   2165: 'FIT417 1 STARBOARD TANK USD FLOW HIGH', class Tank Control Warnings, trigger "2062_Warning_Data_BTCS_WARNING_WORD_03" bit 5
   2166: 'FIT418 3 PORT TANK USD FLOW LOW', class Tank Control Warnings, trigger "2062_Warning_Data_BTCS_WARNING_WORD_03" bit 6
   2164: 'FIT417 1 STARBOARD TANK USD FLOW LOW', class Tank Control Warnings, trigger "2062_Warning_Data_BTCS_WARNING_WORD_03" bit 4
   2162: 'FIT418 1 PORT TANK USD FLOW LOW', class Tank Control Warnings, trigger "2062_Warning_Data_BTCS_WARNING_WORD_03" bit 2
   2163: 'FIT418 1 PORT TANK USD FLOW HIGH', class Tank Control Warnings, trigger "2062_Warning_Data_BTCS_WARNING_WORD_03" bit 3
   2241: 'LS425 5 PORT TANK LEVEL HIGH HIGH', class Tank Control Warnings, trigger "2062_Warning_Data_BTCS_WARNING_WORD_08" bit 1
   2242: 'LS425 5 STARBOARD TANK LEVEL HIGH HIGH', class Tank Control Warnings, trigger "2062_Warning_Data_BTCS_WARNING_WORD_08" bit 2
   2240: 'LS425 4 STARBOARD TANK LEVEL HIGH HIGH', class Tank Control Warnings, trigger "2062_Warning_Data_BTCS_WARNING_WORD_08" bit 0
   2302: 'TT426 1S BWT TEMP HIGH', class Tank Control Warnings, trigger "2062_Warning_Data_BTCS_WARNING_WORD_11" bit 14
   2303: 'TT426 2P BWT TEMP HIGH', class Tank Control Warnings, trigger "2062_Warning_Data_BTCS_WARNING_WORD_11" bit 15
   2243: 'LS425 6 PORT TANK LEVEL HIGH HIGH', class Tank Control Warnings, trigger "2062_Warning_Data_BTCS_WARNING_WORD_08" bit 3
   2247: 'LS425 FP TANK LEVEL HIGH HIGH', class Tank Control Warnings, trigger "2062_Warning_Data_BTCS_WARNING_WORD_08" bit 7
   2248: 'PT415 RIO7 DECK IG PRESSURE LOW', class Tank Control Warnings, trigger "2062_Warning_Data_BTCS_WARNING_WORD_08" bit 8
   2246: 'BTCS_WARNING_WORD_08_BIT_14', class Tank Control Warnings, trigger "2062_Warning_Data_BTCS_WARNING_WORD_08" bit 6
   2244: 'LS425 6 STARBOARD TANK LEVEL HIGH HIGH', class Tank Control Warnings, trigger "2062_Warning_Data_BTCS_WARNING_WORD_08" bit 4
   2245: 'LS425 AP TANK LEVEL HIGH HIGH', class Tank Control Warnings, trigger "2062_Warning_Data_BTCS_WARNING_WORD_08" bit 5
   2234: 'PIT424 RIO1 TANK PRESSURE LOW', class Tank Control Warnings, trigger "2062_Warning_Data_BTCS_WARNING_WORD_07" bit 10
   2235: 'PIT424 RIO1 TANK PRESSURE HIGH', class Tank Control Warnings, trigger "2062_Warning_Data_BTCS_WARNING_WORD_07" bit 11
   2299: 'LT422 APT TANK LEVEL LOW', class Tank Control Warnings, trigger "2062_Warning_Data_BTCS_WARNING_WORD_11" bit 11
   2232: 'PT415 RIO6 DECK IG PRESSURE LOW', class Tank Control Warnings, trigger "2062_Warning_Data_BTCS_WARNING_WORD_07" bit 8
   2233: 'PT415 RIO6 DECK IG PRESSURE HIGH', class Tank Control Warnings, trigger "2062_Warning_Data_BTCS_WARNING_WORD_07" bit 9
   2300: 'TT426 FPT BWT TEMP HIGH', class Tank Control Warnings, trigger "2062_Warning_Data_BTCS_WARNING_WORD_11" bit 12
   2238: 'PIT424 RIO4 TANK PRESSURE LOW', class Tank Control Warnings, trigger "2062_Warning_Data_BTCS_WARNING_WORD_07" bit 14
   2239: 'PIT424 RIO4 TANK PRESSURE HIGH', class Tank Control Warnings, trigger "2062_Warning_Data_BTCS_WARNING_WORD_07" bit 15
   2301: 'TT426 1P BWT TEMP HIGH', class Tank Control Warnings, trigger "2062_Warning_Data_BTCS_WARNING_WORD_11" bit 13
   2236: 'PIT424 RIO3 TANK PRESSURE LOW', class Tank Control Warnings, trigger "2062_Warning_Data_BTCS_WARNING_WORD_07" bit 12
   2237: 'PIT424 RIO3 TANK PRESSURE HIGH', class Tank Control Warnings, trigger "2062_Warning_Data_BTCS_WARNING_WORD_07" bit 13
   2249: 'PT415 RIO7 DECK IG PRESSURE HIGH', class Tank Control Warnings, trigger "2062_Warning_Data_BTCS_WARNING_WORD_08" bit 9
   2264: 'PS436 RIO1 TANK GROUP PRESURE HIGH HIGH', class Tank Control Warnings, trigger "2062_Warning_Data_BTCS_WARNING_WORD_09" bit 8
   2265: 'PS436 RIO2 TANK GROUP PRESURE HIGH HIGH', class Tank Control Warnings, trigger "2062_Warning_Data_BTCS_WARNING_WORD_09" bit 9
   2263: 'LT422 2 PORT TANK LEVEL LOW', class Tank Control Warnings, trigger "2062_Warning_Data_BTCS_WARNING_WORD_09" bit 7
   2261: 'LT422 1 STARBOARD TANK LEVEL LOW', class Tank Control Warnings, trigger "2062_Warning_Data_BTCS_WARNING_WORD_09" bit 5
   2262: 'LT422 2 PORT TANK LEVEL HIGH', class Tank Control Warnings, trigger "2062_Warning_Data_BTCS_WARNING_WORD_09" bit 6
   2266: 'PS436 RIO3 TANK GROUP PRESURE HIGH HIGH', class Tank Control Warnings, trigger "2062_Warning_Data_BTCS_WARNING_WORD_09" bit 10
   2270: 'PS436 RIO7 TANK GROUP PRESURE HIGH HIGH', class Tank Control Warnings, trigger "2062_Warning_Data_BTCS_WARNING_WORD_09" bit 14
   2271: 'LS425 1 PORT TANK LEVEL HIGH HIGH', class Tank Control Warnings, trigger "2062_Warning_Data_BTCS_WARNING_WORD_09" bit 15
   2269: 'PS436 RIO6 TANK GROUP PRESURE HIGH HIGH', class Tank Control Warnings, trigger "2062_Warning_Data_BTCS_WARNING_WORD_09" bit 13
   2267: 'PS436 RIO4 TANK GROUP PRESURE HIGH HIGH', class Tank Control Warnings, trigger "2062_Warning_Data_BTCS_WARNING_WORD_09" bit 11
   2268: 'PS436 RIO5 TANK GROUP PRESURE HIGH HIGH', class Tank Control Warnings, trigger "2062_Warning_Data_BTCS_WARNING_WORD_09" bit 12
   2253: 'LS425 3 PORT TANK LEVEL HIGH HIGH', class Tank Control Warnings, trigger "2062_Warning_Data_BTCS_WARNING_WORD_08" bit 13
   2254: 'LS425 3 STARBOARD TANK LEVEL HIGH HIGH', class Tank Control Warnings, trigger "2062_Warning_Data_BTCS_WARNING_WORD_08" bit 14
   2252: 'LS425 2 STARBOARD TANK LEVEL HIGH HIGH', class Tank Control Warnings, trigger "2062_Warning_Data_BTCS_WARNING_WORD_08" bit 12
   2250: 'LS425 1 STARBOARD TANK LEVEL HIGH HIGH', class Tank Control Warnings, trigger "2062_Warning_Data_BTCS_WARNING_WORD_08" bit 10
   2251: 'LS425 2 PORT TANK LEVEL HIGH HIGH', class Tank Control Warnings, trigger "2062_Warning_Data_BTCS_WARNING_WORD_08" bit 11
   2255: 'LS425 4 PORT TANK LEVEL HIGH HIGH', class Tank Control Warnings, trigger "2062_Warning_Data_BTCS_WARNING_WORD_08" bit 15
   2259: 'LT422 1 PORT TANK LEVEL LOW', class Tank Control Warnings, trigger "2062_Warning_Data_BTCS_WARNING_WORD_09" bit 3
   2260: 'LT422 1 STARBOARD TANK LEVEL HIGH', class Tank Control Warnings, trigger "2062_Warning_Data_BTCS_WARNING_WORD_09" bit 4
   2258: 'LT422 1 PORT TANK LEVEL HIGH', class Tank Control Warnings, trigger "2062_Warning_Data_BTCS_WARNING_WORD_09" bit 2
   2256: 'LT422 FPT TANK LEVEL HIGH', class Tank Control Warnings, trigger "2062_Warning_Data_BTCS_WARNING_WORD_09" bit 0
   2257: 'LT422 FPT TANK LEVEL LOW', class Tank Control Warnings, trigger "2062_Warning_Data_BTCS_WARNING_WORD_09" bit 1
   2298: 'LT422 APT TANK LEVEL HIGH', class Tank Control Warnings, trigger "2062_Warning_Data_BTCS_WARNING_WORD_11" bit 10
   2211: 'PT415 RIO3 DECK IG PRESSURE HIGH', class Tank Control Warnings, trigger "2062_Warning_Data_BTCS_WARNING_WORD_06" bit 3
   2212: 'PT415 RIO4 DECK IG PRESSURE LOW', class Tank Control Warnings, trigger "2062_Warning_Data_BTCS_WARNING_WORD_06" bit 4
   2210: 'PT415 RIO3 DECK IG PRESSURE LOW', class Tank Control Warnings, trigger "2062_Warning_Data_BTCS_WARNING_WORD_06" bit 2
   2208: 'PT415 RIO1 DECK IG PRESSURE LOW', class Tank Control Warnings, trigger "2062_Warning_Data_BTCS_WARNING_WORD_06" bit 0
   2209: 'PT415 RIO1 DECK IG PRESSURE HIGH', class Tank Control Warnings, trigger "2062_Warning_Data_BTCS_WARNING_WORD_06" bit 1
   2213: 'PT415 RIO4 DECK IG PRESSURE HIGH', class Tank Control Warnings, trigger "2062_Warning_Data_BTCS_WARNING_WORD_06" bit 5
   2289: 'TT426 3P BWT TEMP HIGH', class Tank Control Warnings, trigger "2062_Warning_Data_BTCS_WARNING_WORD_11" bit 1
   2216: 'FIT419 5 STARBOARD MBG FLOW LOW', class Tank Control Warnings, trigger "2062_Warning_Data_BTCS_WARNING_WORD_06" bit 8
   2215: 'PT415 RIO5 DECK IG PRESSURE HIGH', class Tank Control Warnings, trigger "2062_Warning_Data_BTCS_WARNING_WORD_06" bit 7
   2288: 'TT426 2S BWT TEMP HIGH', class Tank Control Warnings, trigger "2062_Warning_Data_BTCS_WARNING_WORD_11" bit 0
   2214: 'PT415 RIO5 DECK IG PRESSURE LOW', class Tank Control Warnings, trigger "2062_Warning_Data_BTCS_WARNING_WORD_06" bit 6
   2202: 'FIT420 1 PORT MBG FLOW LOW', class Tank Control Warnings, trigger "2062_Warning_Data_BTCS_WARNING_WORD_05" bit 10
   2203: 'FIT420 1 PORT MBG FLOW HIGH', class Tank Control Warnings, trigger "2062_Warning_Data_BTCS_WARNING_WORD_05" bit 11
   2285: 'LT422 3 STARBOARD TANK LEVEL LOW', class Tank Control Warnings, trigger "2062_Warning_Data_BTCS_WARNING_WORD_10" bit 13
   2200: 'FIT420 1 FPT MBG FLOW LOW', class Tank Control Warnings, trigger "2062_Warning_Data_BTCS_WARNING_WORD_05" bit 8
   2201: 'FIT420 1 FPT MBG FLOW HIGH', class Tank Control Warnings, trigger "2062_Warning_Data_BTCS_WARNING_WORD_05" bit 9
   2286: 'LT422 4 PORT TANK LEVEL HIGH', class Tank Control Warnings, trigger "2062_Warning_Data_BTCS_WARNING_WORD_10" bit 14
   2206: 'FIT420 3 PORT MBG FLOW LOW', class Tank Control Warnings, trigger "2062_Warning_Data_BTCS_WARNING_WORD_05" bit 14
   2207: 'FIT420 3 PORT MBG FLOW HIGH', class Tank Control Warnings, trigger "2062_Warning_Data_BTCS_WARNING_WORD_05" bit 15
   2287: 'LT422 4 PORT TANK LEVEL LOW', class Tank Control Warnings, trigger "2062_Warning_Data_BTCS_WARNING_WORD_10" bit 15
   2204: 'FIT419 1 STARBOARD MBG FLOW LOW', class Tank Control Warnings, trigger "2062_Warning_Data_BTCS_WARNING_WORD_05" bit 12
   2205: 'FIT419 1 STARBOARD MBG FLOW HIGH', class Tank Control Warnings, trigger "2062_Warning_Data_BTCS_WARNING_WORD_05" bit 13
   2217: 'FIT419 5 STARBOARD MBG FLOW HIGH', class Tank Control Warnings, trigger "2062_Warning_Data_BTCS_WARNING_WORD_06" bit 9
   2226: 'PIT424 RIO6 TANK PRESSURE LOW', class Tank Control Warnings, trigger "2062_Warning_Data_BTCS_WARNING_WORD_07" bit 2
   2227: 'PIT424 RIO6 TANK PRESSURE HIGH', class Tank Control Warnings, trigger "2062_Warning_Data_BTCS_WARNING_WORD_07" bit 3
   2295: 'TT426 6P BWT TEMP HIGH', class Tank Control Warnings, trigger "2062_Warning_Data_BTCS_WARNING_WORD_11" bit 7
   2224: 'PIT424 RIO5 TANK PRESSURE LOW', class Tank Control Warnings, trigger "2062_Warning_Data_BTCS_WARNING_WORD_07" bit 0
   2225: 'PIT424 RIO5 TANK PRESSURE HIGH', class Tank Control Warnings, trigger "2062_Warning_Data_BTCS_WARNING_WORD_07" bit 1
   2296: 'LT422 6S TANK LEVEL HIGH', class Tank Control Warnings, trigger "2062_Warning_Data_BTCS_WARNING_WORD_11" bit 8
   2230: 'BTCS_WARNING_WORD_07_BIT_14', class Tank Control Warnings, trigger "2062_Warning_Data_BTCS_WARNING_WORD_07" bit 6
   2231: 'BTCS_WARNING_WORD_07_BIT_15', class Tank Control Warnings, trigger "2062_Warning_Data_BTCS_WARNING_WORD_07" bit 7
   2297: 'LT422 6S TANK LEVEL LOW', class Tank Control Warnings, trigger "2062_Warning_Data_BTCS_WARNING_WORD_11" bit 9
   2228: 'PIT424 RIO7 TANK PRESSURE LOW', class Tank Control Warnings, trigger "2062_Warning_Data_BTCS_WARNING_WORD_07" bit 4
   2229: 'PIT424 RIO7 TANK PRESSURE HIGH', class Tank Control Warnings, trigger "2062_Warning_Data_BTCS_WARNING_WORD_07" bit 5
   2291: 'TT426 4P BWT TEMP HIGH', class Tank Control Warnings, trigger "2062_Warning_Data_BTCS_WARNING_WORD_11" bit 3
   2220: 'FIT419 6 STARBOARD MBG FLOW LOW', class Tank Control Warnings, trigger "2062_Warning_Data_BTCS_WARNING_WORD_06" bit 12
   2219: 'FIT420 6 PORT MBG FLOW HIGH', class Tank Control Warnings, trigger "2062_Warning_Data_BTCS_WARNING_WORD_06" bit 11
   2290: 'TT426 3S BWT TEMP HIGH', class Tank Control Warnings, trigger "2062_Warning_Data_BTCS_WARNING_WORD_11" bit 2
   2218: 'FIT420 6 PORT MBG FLOW LOW', class Tank Control Warnings, trigger "2062_Warning_Data_BTCS_WARNING_WORD_06" bit 10
   2221: 'FIT419 6 STARBOARD MBG FLOW HIGH', class Tank Control Warnings, trigger "2062_Warning_Data_BTCS_WARNING_WORD_06" bit 13
   2293: 'TT426 5P BWT TEMP HIGH', class Tank Control Warnings, trigger "2062_Warning_Data_BTCS_WARNING_WORD_11" bit 5
   2294: 'TT426 5S BWT TEMP HIGH', class Tank Control Warnings, trigger "2062_Warning_Data_BTCS_WARNING_WORD_11" bit 6
   2223: 'FIT420 7 APT MBG FLOW HIGH', class Tank Control Warnings, trigger "2062_Warning_Data_BTCS_WARNING_WORD_06" bit 15
   2292: 'TT426 4S BWT TEMP HIGH', class Tank Control Warnings, trigger "2062_Warning_Data_BTCS_WARNING_WORD_11" bit 4
   2222: 'FIT420 7 APT MBG FLOW LOW', class Tank Control Warnings, trigger "2062_Warning_Data_BTCS_WARNING_WORD_06" bit 14
   2057: 'PT415 RIO5 DECK IG PRESSURE HGH HIGH', class Tank Control Alarms, trigger "2060_Alarm_Data_BTCS_ALARM_WORD_04" bit 9
   2064: 'CV422 3 PORT GAS to TANK VALVE FAULT', class Tank Control Alarms, trigger "2060_Alarm_Data_BTCS_ALARM_WORD_02" bit 3
   2065: 'CV421 1 STARBOARD GAS to TANK VALVE FAULT', class Tank Control Alarms, trigger "2060_Alarm_Data_BTCS_ALARM_WORD_02" bit 2
   2066: 'CV421 3 STARBOARD GAS to TANK VALVE FAULT', class Tank Control Alarms, trigger "2060_Alarm_Data_BTCS_ALARM_WORD_02" bit 4
   2067: 'CV422 5 PORT GAS to TANK VALVE FAULT', class Tank Control Alarms, trigger "2060_Alarm_Data_BTCS_ALARM_WORD_02" bit 7
   2068: 'CV421 4 STARBOARD GAS to TANK VALVE FAULT', class Tank Control Alarms, trigger "2060_Alarm_Data_BTCS_ALARM_WORD_02" bit 6
   2069: 'CV422 4 PORT GAS to TANK VALVE FAULT', class Tank Control Alarms, trigger "2060_Alarm_Data_BTCS_ALARM_WORD_02" bit 5
   2070: 'PS-436 2 BALLAST TANK PRESSURE - HIGH', class Tank Control Alarms, trigger "2060_Alarm_Data_BTCS_ALARM_WORD_01" bit 14
   2071: 'LS-425 2 STARBOARD LEVEL - HIGH HIGH', class Tank Control Alarms, trigger "2060_Alarm_Data_BTCS_ALARM_WORD_01" bit 13
   2072: 'LS-425 2 PORT LEVEL - HIGH HIGH', class Tank Control Alarms, trigger "2060_Alarm_Data_BTCS_ALARM_WORD_01" bit 12
   2073: '600-TX-433 APT O2 MONITOR - LOW', class Tank Control Alarms, trigger "2060_Alarm_Data_BTCS_ALARM_WORD_01" bit 15
   2074: 'CV422 1 PORT GAS to TANK VALVE FAULT', class Tank Control Alarms, trigger "2060_Alarm_Data_BTCS_ALARM_WORD_02" bit 1
   2075: 'CV422 FPT GAS to TANK VALVE FAULT', class Tank Control Alarms, trigger "2060_Alarm_Data_BTCS_ALARM_WORD_02" bit 0
   2076: 'PIT-424 2 STARBOARD TANK PRESSURE - HIGH HIGH', class Tank Control Alarms, trigger "2060_Alarm_Data_BTCS_ALARM_WORD_02" bit 15
   2077: 'PIT-424 2 STARBOARD TANK PRESSURE - LOW LOW', class Tank Control Alarms, trigger "2060_Alarm_Data_BTCS_ALARM_WORD_02" bit 14
   2078: 'PIT-415 2 STARBOARD DECK IG PRESSURE - LOW LOW', class Tank Control Alarms, trigger "2060_Alarm_Data_BTCS_ALARM_WORD_02" bit 10
   2079: 'PIT-415 2 PORT DECK IG PRESSURE - HIGH HIGH', class Tank Control Alarms, trigger "2060_Alarm_Data_BTCS_ALARM_WORD_02" bit 9
   2080: 'PIT-415 2 PORT DECK IG PRESSURE - LOW LOW', class Tank Control Alarms, trigger "2060_Alarm_Data_BTCS_ALARM_WORD_02" bit 8
   2081: 'PIT-415 2 STARBOARD DECK IG PRESSURE - HIGH HIGH', class Tank Control Alarms, trigger "2060_Alarm_Data_BTCS_ALARM_WORD_02" bit 11
   2082: 'PIT-424 2 PORT TANK PRESSURE - HIGH HIGH', class Tank Control Alarms, trigger "2060_Alarm_Data_BTCS_ALARM_WORD_02" bit 13
   2083: 'PIT-424 2 PORT TANK PRESSURE - LOW LOW', class Tank Control Alarms, trigger "2060_Alarm_Data_BTCS_ALARM_WORD_02" bit 12
   2084: 'FIT-418 2 PORT USD FLOW - LOW LOW', class Tank Control Alarms, trigger "2060_Alarm_Data_BTCS_ALARM_WORD_01" bit 0
   2085: 'CV-442 2 PORT GAS to TANK VALVE FAULT', class Tank Control Alarms, trigger "2060_Alarm_Data_BTCS_ALARM_WORD_01" bit 8
   2086: 'FIT-419 2 STARBOARD MBG FLOW - HIGH HIGH', class Tank Control Alarms, trigger "2060_Alarm_Data_BTCS_ALARM_WORD_01" bit 7
   2087: 'CV-441 2 STARBOARD GAS to TANK VALVE FAULT', class Tank Control Alarms, trigger "2060_Alarm_Data_BTCS_ALARM_WORD_01" bit 9
   2088: 'TIT-436 2 STARBOARD BWT TEMP - HIGH HIGH', class Tank Control Alarms, trigger "2060_Alarm_Data_BTCS_ALARM_WORD_01" bit 11
   2089: 'TIT-436 2 PORT BWT TEMP - HIGH HIGH', class Tank Control Alarms, trigger "2060_Alarm_Data_BTCS_ALARM_WORD_01" bit 10
   2090: 'FIT-419 2 STARBOARD MBG FLOW - LOW LOW', class Tank Control Alarms, trigger "2060_Alarm_Data_BTCS_ALARM_WORD_01" bit 6
   2091: 'FIT-420 2 PORT MBG FLOW - HIGH HIGH', class Tank Control Alarms, trigger "2060_Alarm_Data_BTCS_ALARM_WORD_01" bit 3
   2092: 'FIT-420 2 PORT MBG FLOW - LOW LOW', class Tank Control Alarms, trigger "2060_Alarm_Data_BTCS_ALARM_WORD_01" bit 2
   2093: 'FIT-418 2 PORT USD FLOW - HIGH HIGH', class Tank Control Alarms, trigger "2060_Alarm_Data_BTCS_ALARM_WORD_01" bit 1
   2094: 'FIT-417 2 STARBOARD USD FLOW - HIGH HIGH', class Tank Control Alarms, trigger "2060_Alarm_Data_BTCS_ALARM_WORD_01" bit 5
   2095: 'FIT-417 2 STARBOARD USD FLOW - LOW LOW', class Tank Control Alarms, trigger "2060_Alarm_Data_BTCS_ALARM_WORD_01" bit 4
   2040: 'CV422 5 STARBOARD GAS to TANK VALVE FAULT', class Tank Control Alarms, trigger "2060_Alarm_Data_BTCS_ALARM_WORD_03" bit 8
   2039: '', class Tank Control Alarms, trigger "2060_Alarm_Data_BTCS_ALARM_WORD_03" bit 7
   2038: 'PT415 RIO4 DECK IG PRESSURE HGH HIGH', class Tank Control Alarms, trigger "2060_Alarm_Data_BTCS_ALARM_WORD_03" bit 6
   2044: '', class Tank Control Alarms, trigger "2060_Alarm_Data_BTCS_ALARM_WORD_03" bit 12
   2045: '', class Tank Control Alarms, trigger "2060_Alarm_Data_BTCS_ALARM_WORD_03" bit 13
   2043: 'CV422 APT GAS to TANK VALVE FAULT', class Tank Control Alarms, trigger "2060_Alarm_Data_BTCS_ALARM_WORD_03" bit 11
   2041: 'CV422 6 PORT GAS to TANK VALVE FAULT', class Tank Control Alarms, trigger "2060_Alarm_Data_BTCS_ALARM_WORD_03" bit 9
   2042: 'CV422 6 STARBOARD GAS to TANK VALVE FAULT', class Tank Control Alarms, trigger "2060_Alarm_Data_BTCS_ALARM_WORD_03" bit 10
   2037: 'PT415 RIO4 DECK IG PRESSURE LOW LOW', class Tank Control Alarms, trigger "2060_Alarm_Data_BTCS_ALARM_WORD_03" bit 5
   2035: 'PT415 RIO3 DECK IG PRESSURE LOW LOW', class Tank Control Alarms, trigger "2060_Alarm_Data_BTCS_ALARM_WORD_03" bit 3
   2034: 'PT415 RIO1 DECK IG PRESSURE HGH HIGH', class Tank Control Alarms, trigger "2060_Alarm_Data_BTCS_ALARM_WORD_03" bit 2
   2033: '', class Tank Control Alarms, trigger "2060_Alarm_Data_BTCS_ALARM_WORD_03" bit 1
   2032: 'PT415 RIO1 DECK IG PRESSURE LOW LOW', class Tank Control Alarms, trigger "2060_Alarm_Data_BTCS_ALARM_WORD_03" bit 0
   2036: 'PT415 RIO3 DECK IG PRESSURE HGH HIGH', class Tank Control Alarms, trigger "2060_Alarm_Data_BTCS_ALARM_WORD_03" bit 4
   2046: '', class Tank Control Alarms, trigger "2060_Alarm_Data_BTCS_ALARM_WORD_03" bit 14
   2055: '', class Tank Control Alarms, trigger "2060_Alarm_Data_BTCS_ALARM_WORD_04" bit 7
   2056: 'PT415 RIO5 DECK IG PRESSURE LOW LOW', class Tank Control Alarms, trigger "2060_Alarm_Data_BTCS_ALARM_WORD_04" bit 8
   2052: '', class Tank Control Alarms, trigger "2060_Alarm_Data_BTCS_ALARM_WORD_04" bit 4
   2053: '', class Tank Control Alarms, trigger "2060_Alarm_Data_BTCS_ALARM_WORD_04" bit 5
   2054: '', class Tank Control Alarms, trigger "2060_Alarm_Data_BTCS_ALARM_WORD_04" bit 6
   2051: '', class Tank Control Alarms, trigger "2060_Alarm_Data_BTCS_ALARM_WORD_04" bit 3
   2048: '', class Tank Control Alarms, trigger "2060_Alarm_Data_BTCS_ALARM_WORD_04" bit 0
   2047: '', class Tank Control Alarms, trigger "2060_Alarm_Data_BTCS_ALARM_WORD_03" bit 15
   2050: '', class Tank Control Alarms, trigger "2060_Alarm_Data_BTCS_ALARM_WORD_04" bit 2
   2049: '', class Tank Control Alarms, trigger "2060_Alarm_Data_BTCS_ALARM_WORD_04" bit 1
   2159: 'PIT-424 2 STARBOARD TANK PRESSURE - HIGH', class Tank Control Warnings, trigger "2062_Warning_Data_BTCS_WARNING_WORD_02" bit 15
   2157: 'PIT-424 2 PORT TANK PRESSURE - HIGH', class Tank Control Warnings, trigger "2062_Warning_Data_BTCS_WARNING_WORD_02" bit 13
   2132: 'FIT-417 2 STARBOARD USD FLOW - LOW', class Tank Control Warnings, trigger "2062_Warning_Data_BTCS_WARNING_WORD_01" bit 4
   2133: 'FIT-417 2 STARBOARD USD FLOW - HIGH', class Tank Control Warnings, trigger "2062_Warning_Data_BTCS_WARNING_WORD_01" bit 5
   2134: 'FIT-419 2 STARBOARD MBG FLOW - LOW', class Tank Control Warnings, trigger "2062_Warning_Data_BTCS_WARNING_WORD_01" bit 6
   2135: 'FIT-419 2 STARBOARD MBG FLOW - HIGH', class Tank Control Warnings, trigger "2062_Warning_Data_BTCS_WARNING_WORD_01" bit 7
   2136: '600-TX-433 APT O2 MONITOR - LOW', class Tank Control Warnings, trigger "2062_Warning_Data_BTCS_WARNING_WORD_01" bit 8
   2137: '600-TX-433 APT O2 MONITOR - LOW LOW', class Tank Control Warnings, trigger "2062_Warning_Data_BTCS_WARNING_WORD_01" bit 9
   2138: 'TIT-436 2 PORT BWT TEMP - HIGH', class Tank Control Warnings, trigger "2062_Warning_Data_BTCS_WARNING_WORD_01" bit 10
   2139: 'TIT-436 2 STARBOARD BWT TEMP - HIGH', class Tank Control Warnings, trigger "2062_Warning_Data_BTCS_WARNING_WORD_01" bit 11
   2131: 'FIT-420 2 PORT MBG FLOW - HIGH', class Tank Control Warnings, trigger "2062_Warning_Data_BTCS_WARNING_WORD_01" bit 3
   2140: 'BTCS_WARNING_WORD_01_BIT_4', class Tank Control Warnings, trigger "2062_Warning_Data_BTCS_WARNING_WORD_01" bit 12
   2142: 'BTCS_WARNING_WORD_01_BIT_6', class Tank Control Warnings, trigger "2062_Warning_Data_BTCS_WARNING_WORD_01" bit 14
   2143: 'BTCS_WARNING_WORD_01_BIT_7', class Tank Control Warnings, trigger "2062_Warning_Data_BTCS_WARNING_WORD_01" bit 15
   2141: 'BTCS_WARNING_WORD_01_BIT_5', class Tank Control Warnings, trigger "2062_Warning_Data_BTCS_WARNING_WORD_01" bit 13
   2130: 'FIT-420 2 PORT MBG FLOW - LOW', class Tank Control Warnings, trigger "2062_Warning_Data_BTCS_WARNING_WORD_01" bit 2
   2128: 'FIT-418 2 PORT USD FLOW - LOW', class Tank Control Warnings, trigger "2062_Warning_Data_BTCS_WARNING_WORD_01" bit 0
   2129: 'FIT-418 2 PORT USD FLOW - HIGH', class Tank Control Warnings, trigger "2062_Warning_Data_BTCS_WARNING_WORD_01" bit 1
   2158: 'PIT-424 2 STARBOARD TANK PRESSURE - LOW', class Tank Control Warnings, trigger "2062_Warning_Data_BTCS_WARNING_WORD_02" bit 14
   2144: 'TT-426 1 FOR PEACK TANK TEMPERATURE - HIGH', class Tank Control Warnings, trigger "2062_Warning_Data_BTCS_WARNING_WORD_02" bit 0
   2145: 'TT-426 1 PORT TANK TEMPERATURE - HIGH', class Tank Control Warnings, trigger "2062_Warning_Data_BTCS_WARNING_WORD_02" bit 1
   2146: 'TT-426 1 STARBOARD TANK TEMPERATURE - HIGH', class Tank Control Warnings, trigger "2062_Warning_Data_BTCS_WARNING_WORD_02" bit 2
   2147: 'TT-426 3 PORT TANK TEMPERATURE - HIGH', class Tank Control Warnings, trigger "2062_Warning_Data_BTCS_WARNING_WORD_02" bit 3
   2148: 'TT-426 3 STARBOARD TANK TEMPERATURE - HIGH', class Tank Control Warnings, trigger "2062_Warning_Data_BTCS_WARNING_WORD_02" bit 4
   2149: 'TT-426 4 PORT TANK TEMPERATURE - HIGH', class Tank Control Warnings, trigger "2062_Warning_Data_BTCS_WARNING_WORD_02" bit 5
   2150: 'TT-426 4 STARBOARD TANK TEMPERATURE - HIGH', class Tank Control Warnings, trigger "2062_Warning_Data_BTCS_WARNING_WORD_02" bit 6
   2151: 'TT-426 5 PORT TANK TEMPERATURE - HIGH', class Tank Control Warnings, trigger "2062_Warning_Data_BTCS_WARNING_WORD_02" bit 7
   2152: 'PIT-415 2 PORT DECK IG PRESSURE - LOW', class Tank Control Warnings, trigger "2062_Warning_Data_BTCS_WARNING_WORD_02" bit 8
   2153: 'PIT-415 2 PORT DECK IG PRESSURE - HIGH', class Tank Control Warnings, trigger "2062_Warning_Data_BTCS_WARNING_WORD_02" bit 9
   2154: 'PIT-415 2 STARBOARD DECK IG PRESSURE - LOW', class Tank Control Warnings, trigger "2062_Warning_Data_BTCS_WARNING_WORD_02" bit 10
   2155: 'PIT-415 STARBOARD DECK IG PRESSURE - HIGH', class Tank Control Warnings, trigger "2062_Warning_Data_BTCS_WARNING_WORD_02" bit 11
   2156: 'PIT-424 2 PORT TANK PRESSURE - LOW', class Tank Control Warnings, trigger "2062_Warning_Data_BTCS_WARNING_WORD_02" bit 12
   2304: 'FIT417 3S USD OUT OF RANGE', class Tank Control Warnings, trigger "2062_Warning_Data_BTCS_WARNING_WORD_12" bit 0
   2305: 'FIT418 4P USD OUT OF RANGE', class Tank Control Warnings, trigger "2062_Warning_Data_BTCS_WARNING_WORD_12" bit 1
   2306: 'FIT417 4S USD OUT OF RANGE', class Tank Control Warnings, trigger "2062_Warning_Data_BTCS_WARNING_WORD_12" bit 2
   2307: 'FIT418 5P USD OUT OF RANGE', class Tank Control Warnings, trigger "2062_Warning_Data_BTCS_WARNING_WORD_12" bit 3
   2308: 'FIT417 5S USD OUT OF RANGE', class Tank Control Warnings, trigger "2062_Warning_Data_BTCS_WARNING_WORD_12" bit 4
   2309: 'FIT418 6P USD OUT OF RANGE', class Tank Control Warnings, trigger "2062_Warning_Data_BTCS_WARNING_WORD_12" bit 5
   2310: 'FIT417 6S USD OUT OF RANGE', class Tank Control Warnings, trigger "2062_Warning_Data_BTCS_WARNING_WORD_12" bit 6
   2311: 'FIT417 APT USD OUT OF RANGE', class Tank Control Warnings, trigger "2062_Warning_Data_BTCS_WARNING_WORD_12" bit 7
   2312: 'TT426 6S BWT TEMP OUT OF RANGE', class Tank Control Warnings, trigger "2062_Warning_Data_BTCS_WARNING_WORD_12" bit 8
   2313: 'TT426 APT BWT TEMP OUT OF RANGE', class Tank Control Warnings, trigger "2062_Warning_Data_BTCS_WARNING_WORD_12" bit 9
   2314: 'FIT418 FPT USD OUT OF RANGE', class Tank Control Warnings, trigger "2062_Warning_Data_BTCS_WARNING_WORD_12" bit 10
   2315: 'FIT418 1P USD OUT OF RANGE', class Tank Control Warnings, trigger "2062_Warning_Data_BTCS_WARNING_WORD_12" bit 11
   2316: 'FIT417 1S USD OUT OF RANGE', class Tank Control Warnings, trigger "2062_Warning_Data_BTCS_WARNING_WORD_12" bit 12
   2317: 'FIT418 2P USD OUT OF RANGE', class Tank Control Warnings, trigger "2062_Warning_Data_BTCS_WARNING_WORD_12" bit 13
   2318: 'FIT417 2S USD OUT OF RANGE', class Tank Control Warnings, trigger "2062_Warning_Data_BTCS_WARNING_WORD_12" bit 14
   2319: 'FIT418 3P USD OUT OF RANGE', class Tank Control Warnings, trigger "2062_Warning_Data_BTCS_WARNING_WORD_12" bit 15
   2320: 'FIT419 4S MBG FLOW OUT OF RANGE', class Tank Control Warnings, trigger "2062_Warning_Data_BTCS_WARNING_WORD_13" bit 0
   2321: 'FIT420 5P MBG FLOW OUT OF RANGE', class Tank Control Warnings, trigger "2062_Warning_Data_BTCS_WARNING_WORD_13" bit 1
   2322: 'FIT419 5S MBG FLOW OUT OF RANGE', class Tank Control Warnings, trigger "2062_Warning_Data_BTCS_WARNING_WORD_13" bit 2
   2323: 'FIT420 6P MBG FLOW OUT OF RANGE', class Tank Control Warnings, trigger "2062_Warning_Data_BTCS_WARNING_WORD_13" bit 3
   2324: 'FIT419 6S MBG FLOW OUT OF RANGE', class Tank Control Warnings, trigger "2062_Warning_Data_BTCS_WARNING_WORD_13" bit 4
   2325: 'FIT420 APT MBG FLOW OUT OF RANGE', class Tank Control Warnings, trigger "2062_Warning_Data_BTCS_WARNING_WORD_13" bit 5
   2326: 'PT415 RIO1 DECK IG PRESSURE OUT OF RANGE', class Tank Control Warnings, trigger "2062_Warning_Data_BTCS_WARNING_WORD_13" bit 6
   2327: 'PT415 RIO2 DECK IG PRESSURE OUT OF RANGE', class Tank Control Warnings, trigger "2062_Warning_Data_BTCS_WARNING_WORD_13" bit 7
   2328: 'FIT420 FPT MBG FLOW OUT OF RANGE', class Tank Control Warnings, trigger "2062_Warning_Data_BTCS_WARNING_WORD_13" bit 8
   2329: 'FIT420 1P MBG FLOW OUT OF RANGE', class Tank Control Warnings, trigger "2062_Warning_Data_BTCS_WARNING_WORD_13" bit 9
   2330: 'FIT419 1S MBG FLOW OUT OF RANGE', class Tank Control Warnings, trigger "2062_Warning_Data_BTCS_WARNING_WORD_13" bit 10
   2331: 'FIT420 2P MBG FLOW OUT OF RANGE', class Tank Control Warnings, trigger "2062_Warning_Data_BTCS_WARNING_WORD_13" bit 11
   2332: 'FIT419 2S MBG FLOW OUT OF RANGE', class Tank Control Warnings, trigger "2062_Warning_Data_BTCS_WARNING_WORD_13" bit 12
   2333: 'FIT420 3P MBG FLOW OUT OF RANGE', class Tank Control Warnings, trigger "2062_Warning_Data_BTCS_WARNING_WORD_13" bit 13
   2334: 'FIT419 3S MBG FLOW OUT OF RANGE', class Tank Control Warnings, trigger "2062_Warning_Data_BTCS_WARNING_WORD_13" bit 14
   2335: 'FIT420 4P MBG FLOW OUT OF RANGE', class Tank Control Warnings, trigger "2062_Warning_Data_BTCS_WARNING_WORD_13" bit 15
   2336: 'PIT424 RIO4 TANK PRESSURE OUT OF RANGE', class Tank Control Warnings, trigger "2062_Warning_Data_BTCS_WARNING_WORD_14" bit 0
   2337: 'PIT424 RIO5 TANK PRESSURE OUT OF RANGE', class Tank Control Warnings, trigger "2062_Warning_Data_BTCS_WARNING_WORD_14" bit 1
   2338: 'PIT424 RIO6 TANK PRESSURE OUT OF RANGE', class Tank Control Warnings, trigger "2062_Warning_Data_BTCS_WARNING_WORD_14" bit 2
   2339: 'PIT424 RIO7 TANK PRESSURE OUT OF RANGE', class Tank Control Warnings, trigger "2062_Warning_Data_BTCS_WARNING_WORD_14" bit 3
   2340: 'LT422 FPT TANK LEVEL OUT OF RANGE', class Tank Control Warnings, trigger "2062_Warning_Data_BTCS_WARNING_WORD_14" bit 4
   2341: 'LT422 1P TANK LEVEL OUT OF RANGE', class Tank Control Warnings, trigger "2062_Warning_Data_BTCS_WARNING_WORD_14" bit 5
   2342: 'LT422 1S TANK LEVEL OUT OF RANGE', class Tank Control Warnings, trigger "2062_Warning_Data_BTCS_WARNING_WORD_14" bit 6
   2343: 'LT422 2P TANK LEVEL OUT OF RANGE', class Tank Control Warnings, trigger "2062_Warning_Data_BTCS_WARNING_WORD_14" bit 7
   2344: 'PT415 RIO3 DECK IG PRESSURE OUT OF RANGE', class Tank Control Warnings, trigger "2062_Warning_Data_BTCS_WARNING_WORD_14" bit 8
   2345: 'PT415 RIO4 DECK IG PRESSURE OUT OF RANGE', class Tank Control Warnings, trigger "2062_Warning_Data_BTCS_WARNING_WORD_14" bit 9
   2346: 'PT415 RIO5 DECK IG PRESSURE OUT OF RANGE', class Tank Control Warnings, trigger "2062_Warning_Data_BTCS_WARNING_WORD_14" bit 10
   2347: 'PT415 RIO6 DECK IG PRESSURE OUT OF RANGE', class Tank Control Warnings, trigger "2062_Warning_Data_BTCS_WARNING_WORD_14" bit 11
   2348: 'PT415 RIO7 DECK IG PRESSURE OUT OF RANGE', class Tank Control Warnings, trigger "2062_Warning_Data_BTCS_WARNING_WORD_14" bit 12
   2349: 'PIT424 RIO1 TANK PRESSURE OUT OF RANGE', class Tank Control Warnings, trigger "2062_Warning_Data_BTCS_WARNING_WORD_14" bit 13
   2350: 'PIT424 RIO2 TANK PRESSURE OUT OF RANGE', class Tank Control Warnings, trigger "2062_Warning_Data_BTCS_WARNING_WORD_14" bit 14
   2351: 'PIT424 RIO3 TANK PRESSURE OUT OF RANGE', class Tank Control Warnings, trigger "2062_Warning_Data_BTCS_WARNING_WORD_14" bit 15
   2352: 'LT422 6S TANK LEVEL OUT OF RANGE', class Tank Control Warnings, trigger "2062_Warning_Data_BTCS_WARNING_WORD_15" bit 0
   2353: 'LT422 APT TANK LEVEL OUT OF RANGE', class Tank Control Warnings, trigger "2062_Warning_Data_BTCS_WARNING_WORD_15" bit 1
   2354: '600-TX-433 APT O2 MONITOR OUT OF RANGE', class Tank Control Warnings, trigger "2062_Warning_Data_BTCS_WARNING_WORD_15" bit 2
   2355: 'PH426 FPT OUT OF RANGE', class Tank Control Warnings, trigger "2062_Warning_Data_BTCS_WARNING_WORD_15" bit 3
   2356: 'PH426 1P OUT OF RANGE', class Tank Control Warnings, trigger "2062_Warning_Data_BTCS_WARNING_WORD_15" bit 4
   2357: 'PH426 1S OUT OF RANGE', class Tank Control Warnings, trigger "2062_Warning_Data_BTCS_WARNING_WORD_15" bit 5
   2358: 'PH426 2P OUT OF RANGE', class Tank Control Warnings, trigger "2062_Warning_Data_BTCS_WARNING_WORD_15" bit 6
   2359: 'PH426 2S OUT OF RANGE', class Tank Control Warnings, trigger "2062_Warning_Data_BTCS_WARNING_WORD_15" bit 7
   2360: 'LT422 2S TANK LEVEL OUT OF RANGE', class Tank Control Warnings, trigger "2062_Warning_Data_BTCS_WARNING_WORD_15" bit 8
   2361: 'LT422 3P TANK LEVEL OUT OF RANGE', class Tank Control Warnings, trigger "2062_Warning_Data_BTCS_WARNING_WORD_15" bit 9
   2362: 'LT422 3S TANK LEVEL OUT OF RANGE', class Tank Control Warnings, trigger "2062_Warning_Data_BTCS_WARNING_WORD_15" bit 10
   2363: 'LT422 4P TANK LEVEL OUT OF RANGE', class Tank Control Warnings, trigger "2062_Warning_Data_BTCS_WARNING_WORD_15" bit 11
   2364: 'LT422 4S TANK LEVEL OUT OF RANGE', class Tank Control Warnings, trigger "2062_Warning_Data_BTCS_WARNING_WORD_15" bit 12
   2365: 'LT422 5P TANK LEVEL OUT OF RANGE', class Tank Control Warnings, trigger "2062_Warning_Data_BTCS_WARNING_WORD_15" bit 13
   2366: 'LT422 5S TANK LEVEL OUT OF RANGE', class Tank Control Warnings, trigger "2062_Warning_Data_BTCS_WARNING_WORD_15" bit 14
   2367: 'LT422 6P TANK LEVEL OUT OF RANGE', class Tank Control Warnings, trigger "2062_Warning_Data_BTCS_WARNING_WORD_15" bit 15
   2368: 'PH425 6S OUT OF RANGE', class Tank Control Warnings, trigger "2062_Warning_Data_BTCS_WARNING_WORD_16" bit 0
   2369: 'PH426 APT OUT OF RANGE', class Tank Control Warnings, trigger "2062_Warning_Data_BTCS_WARNING_WORD_16" bit 1
   2370: 'DO428 FPT OUT OF RANGE', class Tank Control Warnings, trigger "2062_Warning_Data_BTCS_WARNING_WORD_16" bit 2
   2371: 'DO428 1P OUT OF RANGE', class Tank Control Warnings, trigger "2062_Warning_Data_BTCS_WARNING_WORD_16" bit 3
   2372: 'DO427 1S OUT OF RANGE', class Tank Control Warnings, trigger "2062_Warning_Data_BTCS_WARNING_WORD_16" bit 4
   2373: 'DO428 2P OUT OF RANGE', class Tank Control Warnings, trigger "2062_Warning_Data_BTCS_WARNING_WORD_16" bit 5
   2374: 'DO427 2S OUT OF RANGE', class Tank Control Warnings, trigger "2062_Warning_Data_BTCS_WARNING_WORD_16" bit 6